
text list "SDC_G120D": 0 ''; 0 'Antrieb hat keine Störung / kein Fehlercode'; 1000 'Softwarefehler intern'; 1001 'FloatingPoint Ausnahme'; 1002 'Softwarefehler intern'; 1003 'Quittungsverzug bei Speicherzugriff'; 1004 'Softwarefehler intern'; 1005 'Datei Upload/Download fehlgeschlagen'; 1009 'CU: Regelungsbaugruppe Übertemperatur'; 1010 'Antriebstyp unbekannt'; 1015 'Softwarefehler intern'; 1016 'Firmware verändert'; 1017 'Komponentenlisten verändert'; 1018 'Hochlauf mehrmals abgebrochen'; 1019 'Wechselmedium schreiben fehlgeschlagen'; 1020 'RAM disk Schreiben fehlgeschlagen'; 1021 'Wechselmedium als USB-Datenträger von PC verwendet'; 1023 'Software Timeout intern'; 1028 'Konfigurationsfehler'; 1030 'Lebenszeichenausfall bei Steuerungshoheit'; 1033 'Einheitenumschaltung: Bezugsparameterwert ungültig'; 1034 'Einheitenumschaltung: Berechnung Parameterwerte nach Bezugswertänderung fehlgeschlagen'; 1035 'ACX: Parametersicherungsdateien beschädigt'; 1036 'ACX: Parametersicherungsdatei fehlt'; 1038 'ACX: Parametersicherungsdatei laden fehlgeschlagen'; 1039 'ACX: Parametersicherungsdatei schreiben fehlgeschlagen'; 1040 'Parameter sichern und POWER ON erforderlich'; 1042 'Parameterfehler beim Projekt-Download'; 1043 'Schwerer Fehler beim Projekt-Download'; 1044 'CU: Beschreibungsdaten fehlerhaft'; 1045 'Projektierungsdaten ungültig'; 1049 'Schreiben in Datei nicht möglich'; 1054 'CU: Systemgrenze überschritten'; 1064 'CU: Interner Fehler (CRC)'; 1066 'Zwischenspeicher: Füllstand 70 % erreicht oder überschritten'; 1067 'Zwischenspeicher: Füllstand 100 % erreicht'; 1068 'CU: Datenspeicher Speicherüberlauf'; 1069 'Parametersicherung und Gerät inkompatibel'; 1072 'Speicherkarte aus Sicherungskopie wieder hergestellt'; 1073 'POWER ON für Sicherungskopie auf Speicherkarte erforderlich'; 1105 'CU: Speicher nicht ausreichend'; 1107 'Speichern auf Speicherkarte fehlgeschlagen'; 1112 'CU: Leistungsteil unzulässig'; 1120 'Initialisierung Klemmen fehlgeschlagen'; 1122 'Frequenz am Messtastereingang zu hoch'; 1205 'CU: Zeitscheibenüberlauf'; 1250 'CU: CU-EEPROM Read-Only-Daten fehlerhaft'; 1251 'CU: CU-EEPROM Read-Write-Daten fehlerhaft'; 1257 'CU: Firmware-Version veraltet'; 1340 'Topologie: Zu viele Komponenten an einem Strang'; 1505 'BICO: Verschaltung kann nicht hergestellt werden'; 1510 'BICO: Signalquelle ist nicht Float'; 1511 'BICO: Verschaltung mit unterschiedlicher Normierung'; 1512 'BICO: Keine Normierung vorhanden'; 1513 'BICO: Verschaltung DO-übergreifend mit unterschiedlicher Normierung'; 1514 'BICO: Fehler beim Schreiben während Reconnect'; 1515 'BICO: Parameterschreiben nicht erlaubt da Steuerungshoheit aktiv'; 1590 'Antrieb: Motor Wartungsintervall abgelaufen'; 1600 'SI P1: STOP A ausgelöst'; 1611 'SI P1: Defekt in einem Überwachungskanal'; 1620 'SI P1: Sicher abgeschaltetes Moment aktiv'; 1625 'SI P1: Lebenszeichen in Safety-Daten fehlerhaft'; 1649 'SI P1: Softwarefehler intern'; 1650 'SI P1: Abnahmetest erforderlich'; 1651 'SI P1: Synchronisation Safety-Zeitscheiben fehlgeschlagen'; 1653 'SI P1: PROFIBUS/PROFINET-Projektierung fehlerhaft'; 1654 'SI P1: PROFIsafe-Projektierung abweichend'; 1655 'SI P1: Abgleich der Überwachungsfunktionen'; 1656 'SI P1: Parameter Prozessor 2 fehlerhaft'; 1658 'SI P1: PROFIsafe-Telegrammnummer ungeeignet'; 1659 'SI P1: Schreibauftrag für Parameter abgewiesen'; 1660 'SI P1: Sichere Funktionen nicht unterstützt'; 1661 'SI P1: Simulation der Safety Eingänge aktiv'; 1662 'Fehler interne Kommunikation'; 1663 'SI P1: Kopieren der SI-Parameter abgelehnt'; 1665 'SI P1: System ist defekt'; 1666 'SI Motion P1: Statisches 1-Signal am F-DI für sichere Quittierung'; 1669 'SI Motion: Kombination von Motor und Leistungsteil ungünstig'; 1680 'SI Motion P1: Prüfsummenfehler sichere Überwachungen'; 1681 'SI Motion P1: Parameterwert falsch'; 1682 'SI Motion P1: Überwachungsfunktion nicht unterstützt'; 1683 'SI Motion P1: SLS-Freigabe fehlt'; 1690 'SI Motion: Datensicherungsproblem beim NVRAM'; 1692 'SI Motion P1: Parameterwert geberlos unzulässig'; 1693 'SI Motion P1: Safety-Parametrierung geändert POWER ON erforderlich'; 1696 'SI Motion: Testanwahl der Bewegungsüberwachungen im Hochlauf'; 1697 'SI Motion: Test der Bewegungsüberwachungen erforderlich'; 1698 'SI P1: Inbetriebnahmemodus aktiv'; 1699 'SI P1: Test der Abschaltpfade erforderlich'; 1700 'SI Motion P1: STOP A ausgelöst'; 1701 'SI Motion P1: STOP B ausgelöst'; 1706 'SI Motion P1: SAM/SBR Grenze überschritten'; 1711 'SI Motion P1: Defekt in einem Überwachungskanal'; 1712 'SI Motion P1: Defekt bei F-IO-Verarbeitung'; 1714 'SI Motion P1: Sicher begrenzte Geschwindigkeit überschritten'; 1716 'SI Motion P1: Toleranz für sichere Bewegungsrichtung überschritten'; 1770 'SI Motion P1: Diskrepanzfehler der fehlersicheren Eingänge'; 1772 'SI Motion P1: Teststop fehlersichere Eingänge/Ausgänge aktiv'; 1773 'SI Motion P1: Teststop fehlerhaft'; 1774 'SI Motion P1: Teststop notwendig'; 1796 'SI P1: Warten auf Kommunikation'; 1798 'SI Motion P1: Teststop läuft'; 1799 'SI Motion P1: Abnahmetestmodus aktiv'; 1900 'PROFIBUS: Konfigurationstelegramm fehlerhaft'; 1910 'Feldbus SS Sollwert Timeout'; 1920 'PROFIBUS: Unterbrechung zyklische Verbindung'; 1945 'PROFIBUS: Verbindung zum Publisher gestört'; 1946 'PROFIBUS: Verbindung zum Publisher abgebrochen'; 1951 'CU SYNC: Synchronisation Applikationstakt fehlt'; 1953 'CU SYNC: Synchronisation nicht abgeschlossen'; 2050 'Trace: Start nicht möglich'; 2055 'Trace: Aufzeichnungsdauer zu klein'; 2056 'Trace: Aufzeichnungstakt zu klein'; 2057 'Trace: Zeitscheibentakt ungültig'; 2058 'Trace: Zeitscheibentakt für Endlostrace ungültig'; 2059 'Trace: Zeitscheibentakt für 2 x 8 Aufzeichnungskanäle ungültig'; 2060 'Trace: Aufzuzeichnendes Signal fehlt'; 2061 'Trace: Signal ungültig'; 2062 'Trace: Triggersignal ungültig'; 2063 'Trace: Datentyp ungültig'; 2070 'Trace: Parameter nicht änderbar'; 2075 'Trace: Pretriggerzeit zu groß'; 2080 'Trace: Parametrierung wegen Einheitenumschaltung gelöscht'; 2097 'MTrace: Mehrfachtrace aktivieren nicht möglich'; 2098 'MTrace: Speichern nicht möglich'; 2099 'Trace: Speicherplatz der Control Unit nicht ausreichend'; 2150 'OA: Applikation nicht ladbar'; 2151 'OA: Softwarefehler intern'; 2152 'OA: Speicher nicht ausreichend'; 3000 'NVRAM Fehler bei Aktion'; 3001 'NVRAM Prüfsumme fehlerhaft'; 3505 'CU: Analogeingang Drahtbruch'; 3510 'CU: Kalibrierdaten nicht plausibel'; 5000 'Leistungsteil: Übertemperatur Kühlkörper Wechselrichter'; 5001 'Leistungsteil: Übertemperatur Sperrschicht Chip'; 5002 'Leistungsteil: Übertemperatur Zuluft'; 5004 'Leistungsteil: Übertemperatur Gleichrichter'; 5006 'Leistungsteil: Übertemperatur Thermisches Modell'; 6310 'Anschlussspannung (p0210) fehlerhaft parametriert'; 6921 'Bremswiderstand Phasenunsymmetrie'; 6922 'Bremswiderstand Phasenausfall'; 7011 'Antrieb: Motor Übertemperatur'; 7012 'Antrieb: Motortemperaturmodell 1 Übertemperatur'; 7014 'Antrieb: Motortemperaturmodell Konfiguration Warnung'; 7015 'Antrieb: Motortemperatursensor Warnung'; 7016 'Antrieb: Motortemperatursensor Störung'; 7080 'Antrieb: Regelungsparameter fehlerhaft'; 7082 'Makro: Ausführung nicht möglich'; 7083 'Makro: ACX-File nicht gefunden'; 7084 'Makro: Bedingung für WaitUntil nicht erfüllt'; 7086 'Einheitenumschaltung: Parametergrenzverletzung durch Bezugswertänderung'; 7088 'Einheitenumschaltung: Parametergrenzverletzung durch Einheitenumschaltung'; 7089 'Einheitenumschaltung: Funktionsmodul aktivieren ist blockiert weil Einheiten umgeschaltet'; 7200 'Antrieb: Steuerungshoheit EIN-Befehl steht an'; 7220 'Antrieb: Führung durch PLC fehlt'; 7300 'Antrieb: Netzschütz Rückmeldung fehlt'; 7320 'Antrieb: Automatischer Wiederanlauf abgebrochen'; 7321 'Antrieb: Automatischer Wiederanlauf aktiv'; 7330 'Fangen: Gemessener Suchstrom zu klein'; 7331 'Fangen: Funktion nicht unterstützt'; 7400 'Antrieb: Zwischenkreisspannungs-Maximum-Regler aktiv'; 7401 'Antrieb: Zwischenkreisspannungs-Maximum-Regler deaktiviert'; 7402 'Antrieb: Zwischenkreisspannungs-Minimum-Regler aktiv'; 7404 'Antrieb: Zwischenkreisspannungsüberwachnung Vdc_Max'; 7405 'Antrieb: Kinetische Pufferung minimale Drehzahl unterschritten'; 7406 'Antrieb: Kinetische Pufferung maximale Dauer überschritten'; 7409 'Antrieb: U/f-Steuerung Strombegrenzungsregler aktiv'; 7410 'Antrieb: Stromreglerausgang begrenzt'; 7411 'Antrieb: Flussreglerausgang begrenzt'; 7416 'Antrieb: Konfiguration Flussregler'; 7426 'Technologieregler Istwert begrenzt'; 7428 'Technologieregler Parametrierfehler'; 7435 'Antrieb: Hochlaufgebersetzen bei geberloser Vektorregelung'; 7440 'EPOS: Ruckzeit wird begrenzt'; 7441 'LR: Lageoffset der Absolutwertgeberjustage sichern'; 7442 'LR: Multiturn passt nicht zum Modulobereich'; 7443 'LR: Referenzpunkt-Koordinate nicht im zulässigen Bereich'; 7450 'LR: Stillstandsüberwachung hat angesprochen'; 7451 'LR: Positionierüberwachung hat angesprochen'; 7452 'LR: Schleppabstand zu groß'; 7453 'LR: Lageistwertaufbereitung fehlerhaft'; 7454 'LR: Lageistwertaufbereitung hat keinen gültigen Geber'; 7455 'EPOS: Maximalgeschwindigkeit begrenzt'; 7456 'EPOS: Sollgeschwindigkeit begrenzt'; 7457 'EPOS: Eingangssignale Kombination unzulässig'; 7458 'EPOS: Referenznocken nicht gefunden'; 7459 'EPOS: Keine Nullmarke vorhanden'; 7460 'EPOS: Referenznockenende nicht gefunden'; 7461 'EPOS: Referenzpunkt nicht gesetzt'; 7462 'EPOS: Angewählte Verfahrsatznummer existiert nicht'; 7463 'EPOS: Externer Satzwechsel im Verfahrsatz nicht angefordert'; 7464 'EPOS: Verfahrsatz ist inkonsistent'; 7465 'EPOS: Verfahrsatz hat keinen Folgesatz'; 7466 'EPOS: Verfahrsatznummer mehrfach vergeben'; 7467 'EPOS: Verfahrsatz hat unzulässigen Auftragsparameter'; 7468 'EPOS: Verfahrsatz Sprungziel existiert nicht'; 7469 'EPOS: Verfahrsatz Zielposition < Software-Endschalter Minus'; 7470 'EPOS: Verfahrsatz Zielposition > Software-Endschalter Plus'; 7471 'EPOS: Verfahrsatz Zielposition außerhalb Modulobereich'; 7472 'EPOS: Verfahrsatz ABS_POS/ABS_NEG nicht möglich'; 7473 'EPOS: Verfahrbereichsanfang angefahren'; 7474 'EPOS: Verfahrbereichsende angefahren'; 7475 'EPOS: Zielposition < Verfahrbereichsanfang'; 7476 'EPOS: Zielposition > Verfahrbereichsende'; 7477 'EPOS: Zielposition < Software-Endschalter Minus'; 7478 'EPOS: Zielposition > Software-Endschalter Plus'; 7479 'EPOS: Software-Endschalter Minus angefahren'; 7480 'EPOS: Software-Endschalter Plus angefahren'; 7481 'EPOS: Achsposition < Software-Endschalter Minus'; 7482 'EPOS: Achsposition > Software-Endschalter Plus'; 7483 'EPOS: Fahren auf Festanschlag Klemmmoment nicht erreicht'; 7484 'EPOS: Festanschlag außerhalb Überwachungsfenster'; 7485 'EPOS: Festanschlag nicht erreicht'; 7486 'EPOS: Zwischenhalt fehlt'; 7487 'EPOS: Verfahrauftrag verwerfen fehlt'; 7488 'EPOS: Relative Positionierung nicht möglich'; 7489 'EPOS: Referenzpunktkorrektur außerhalb Fenster'; 7490 'EPOS: Freigabe während Verfahren weggenommen'; 7491 'EPOS: STOP-Nocken Minus angefahren'; 7492 'EPOS: STOP-Nocken Plus angefahren'; 7493 'LR: Überlauf des Wertebereiches für Lageistwert'; 7494 'LR: Antriebsdatensatz-Umschaltung während Betrieb'; 7495 'LR: Referenzfunktion abgebrochen'; 7496 'EPOS: Freigabe nicht möglich'; 7497 'LR: Lagesetzwert aktiviert'; 7498 'LR: Messtasterauswertung nicht möglich'; 7499 'EPOS: Umkehrnocken mit falscher Verfahrrichtung angefahren'; 7503 'EPOS: STOP-Nocken mit falscher Verfahrrichtung angefahren'; 7505 'EPOS: Auftrag Festanschlag bei U/f/SLVC-Betrieb nicht möglich'; 7530 'Antrieb: Antriebsdatensatz DDS nicht vorhanden'; 7531 'Antrieb: Befehlsdatensatz CDS nicht vorhanden'; 7550 'Antrieb: Geberparameter zurücksetzen nicht möglich'; 7552 'Antrieb Geber: Geberkonfiguration nicht unterstützt'; 7553 'Antrieb Geber: Sensor Module Konfiguration nicht unterstützt'; 7557 'Geber 1: Referenzpunkt-Koordinate nicht im zulässigen Bereich'; 7558 'Geber 2: Referenzpunkt-Koordinate nicht im zulässigen Bereich'; 7563 'Antrieb Geber: XIST1_ERW Konfiguration fehlerhaft'; 7565 'Antrieb: Geberfehler PROFIdrive-Geberschnittstelle 1'; 7566 'Antrieb: Geberfehler PROFIdrive-Geberschnittstelle 2'; 7577 'Geber 1: Messtasterauswertung nicht möglich'; 7578 'Geber 2: Messtasterauswertung nicht möglich'; 7581 'Geber 1: Lageistwertaufbereitung fehlerhaft'; 7582 'Geber 2: Lageistwertaufbereitung fehlerhaft'; 7584 'Geber 1: Lagesetzwert aktiviert'; 7585 'Geber 2: Lagesetzwert aktiviert'; 7587 'Geber 1: Lageistwertaufbereitung hat keinen gültigen Geber'; 7588 'Geber 2: Lageistwertaufbereitung hat keinen gültigen Geber'; 7590 'Geber 1: Antriebsdatensatz-Umschaltung während Betrieb'; 7591 'Geber 2: Antriebsdatensatz-Umschaltung während Betrieb'; 7593 'Geber 1: Wertebereich für Lageistwert überschritten'; 7594 'Geber 2: Wertebereich für Lageistwert überschritten'; 7596 'Geber 1: Referenzfunktion abgebrochen'; 7597 'Geber 2: Referenzfunktion abgebrochen'; 7599 'Geber 1: Justage nicht möglich'; 7600 'Geber 2: Justage nicht möglich'; 7800 'Antrieb: Kein Leistungsteil vorhanden'; 7801 'Antrieb: Motor Überstrom'; 7802 'Antrieb: Einspeisung oder Leistungsteil nicht bereit'; 7805 'Antrieb: Leistungsteil Überlastung I2t'; 7806 'Antrieb: Generatorische Leistungsgrenze überschritten (F3E)'; 7807 'Antrieb: Kurzschluss/Erdschluss erkannt'; 7808 'HF Damping Module: Dämpfung nicht bereit'; 7810 'Antrieb: Leistungsteil-EEPROM ohne Nenndaten'; 7850 'Externe Warnung 1'; 7851 'Externe Warnung 2'; 7852 'Externe Warnung 3'; 7860 'Externe Störung 1'; 7861 'Externe Störung 2'; 7862 'Externe Störung 3'; 7900 'Antrieb: Motor blockiert'; 7901 'Antrieb: Motor Überdrehzahl'; 7902 'Antrieb: Motor gekippt'; 7903 'Antrieb: Motor Drehzahlabweichung'; 7910 'Antrieb: Motor Übertemperatur'; 7920 'Antrieb: Drehmoment/Drehzahl zu niedrig'; 7921 'Antrieb: Drehmoment/Drehzahl zu hoch'; 7922 'Antrieb: Drehmoment/Drehzahl außerhalb Toleranz'; 7923 'Antrieb: Drehmoment/Drehzahl zu niedrig'; 7924 'Antrieb: Drehmoment/Drehzahl zu hoch'; 7925 'Antrieb: Drehmoment/Drehzahl außerhalb Toleranz'; 7927 'Gleichstrombremsung aktiv'; 7929 'Antrieb: Kein Motor erkannt'; 7936 'Antrieb: Lastausfall'; 7950 'Motorparameter fehlerhaft'; 7967 'Antrieb: Pollageidentifikation interner Fehler'; 7968 'Antrieb: Lq-Ld-Messung fehlerhaft'; 7969 'Antrieb: Pollageidentifikation fehlerhaft'; 7975 'Antrieb: Fahren bis Nullmarke - Sollwertvorgabe erwartet'; 7976 'Antrieb: Geberfeinabgleich aktiviert'; 7980 'Antrieb: Drehende Messung aktiviert'; 7981 'Antrieb: Drehende Messung Freigaben fehlen'; 7983 'Antrieb: Drehende Messung Sättigungskennlinie'; 7984 'Antrieb: Drehzahlregleroptimierung Trägheitsmoment'; 7985 'Antrieb: Drehzahlregleroptimierung (Schwingungstest)'; 7986 'Antrieb: Drehende Messung Hochlaufgeber'; 7988 'Antrieb: Drehende Messung Keine Konfiguration ausgewählt'; 7990 'Antrieb: Motordatenidentifikation fehlerhaft'; 7991 'Antrieb: Motordatenidentifikation aktiviert'; 7994 'Antrieb: Motordatenidentifikation nicht durchgeführt'; 8010 'CU: Analog-Digital-Wandler'; 8501 'PROFINET: Sollwert Timeout'; 8502 'PROFINET: Überwachungszeit Lebenszeichen abgelaufen'; 8511 'PROFINET: Empfangs-Konfigurationsdaten ungültig'; 8526 'PROFINET: Keine zyklische Verbindung'; 8565 'PROFINET: Konsistenzfehler bei Einstellparametern'; 8760 'CAN: Überschreitung maximaler Größe des PZD IF'; 8800 'PROFIenergy Energiesparmodus aktiv'; 8802 'PROFIenergy Inkrementalgeberversorgung ausschalten nicht möglich'; 13009 'Lizenzierung OA-Applikation nicht lizenziert'; 13100 'Know-how-Schutz: Kopierschutzfehler'; 13101 'Know-how-Schutz: Kopierschutz nicht aktivierbar'; 13102 'Know-how-Schutz: Konsistenzfehler der geschützten Daten'; 30001 'Leistungsteil: Überstrom'; 30002 'Leistungsteil: Zwischenkreisspannung Überspannung'; 30003 'Leistungsteil: Zwischenkreisspannung Unterspannung'; 30004 'Leistungsteil: Übertemperatur Kühlkörper Wechselrichter'; 30005 'Leistungsteil: Überlastung I2t'; 30011 'Leistungsteil: Netzphasenausfall im Hauptstromkreis'; 30015 'Leistungsteil: Phasenausfall Motorleitung'; 30016 'Leistungsteil: Lastversorgung ausgeschaltet'; 30017 'Leistungsteil: Hardware Strombegrenzung zu oft angesprochen'; 30021 'Leistungsteil: Erdschluss'; 30022 'Leistungsteil: Überwachung U_ce'; 30024 'Leistungsteil: Übertemperatur Thermisches Modell'; 30025 'Leistungsteil: Übertemperatur Chip'; 30027 'Leistungsteil: Vorladung Zwischenkreis Zeitüberwachung'; 30031 'Leistungsteil: Hardware Strombegrenzung in Phase U'; 30032 'Leistungsteil: Hardware Strombegrenzung in Phase V'; 30033 'Leistungsteil: Hardware Strombegrenzung in Phase W'; 30034 'Leistungsteil: Übertemperatur Innenraum'; 30042 'Leistungsteil: Lüfter hat maximale Betriebsstunden erreicht'; 30052 'EEPROM Daten fehlerhaft'; 30054 'Leistungsteil: Unterspannung bei Bremse öffnen'; 30057 'Leistungsteil: Netzunsymmetrie'; 30071 'Keine neuen Istwerte von Power Module empfangen'; 30072 'Keine Sollwerte mehr an Power Module übertragbar'; 30074 'Kommunikationsfehler zwischen Control Unit und Power Module'; 30080 'Leistungsteil: Stromanstieg zu schnell'; 30081 'Leistungsteil: Schalthandlungen zu häufig'; 30105 'LT: Istwerterfassung fehlerhaft'; 30502 'Leistungsteil: Zwischenkreis Überspannung'; 30600 'SI P2: STOP A ausgelöst'; 30611 'SI P2: Defekt in einem Überwachungskanal'; 30620 'SI P2: Sicher abgeschaltetes Moment aktiv'; 30625 'SI P2: Lebenszeichen in Safety-Daten fehlerhaft'; 30649 'SI P2: Softwarefehler intern'; 30650 'SI P2: Abnahmetest erforderlich'; 30651 'SI P2: Synchronisation mit Control Unit fehlgeschlagen'; 30655 'SI P2: Abgleich der Überwachungsfunktionen'; 30656 'SI P2: Parameter Prozessor 2 fehlerhaft'; 30659 'SI P2: Schreibauftrag für Parameter abgewiesen'; 30662 'Fehler in interner Kommunikation'; 30664 'Fehler in der Hochlaufphase'; 30665 'SI P2: System ist defekt'; 30666 'SI Motion P2: Statisches 1-Signal am F-DI für sichere Quittierung'; 30680 'SI Motion P2: Prüfsummenfehler sichere Überwachungen'; 30681 'SI Motion P2: Parameterwert falsch'; 30682 'SI Motion P2: Überwachungsfunktion nicht unterstützt'; 30683 'SI Motion P2: SLS-Freigabe fehlt'; 30692 'SI Motion P2: Parameterwert falsch geberlos'; 30693 'SI P2: Safety-Parametrierung geändert POWER ON erforderlich'; 30700 'SI Motion P2: STOP A ausgelöst'; 30701 'SI Motion P2: STOP B ausgelöst'; 30706 'SI Motion P2: SAM/SBR Grenze überschritten'; 30711 'SI Motion P2: Defekt in einem Überwachungskanal'; 30712 'SI Motion P2: Defekt bei F-IO-Verarbeitung'; 30714 'SI Motion P2: Sicher begrenzte Geschwindigkeit überschritten'; 30716 'SI Motion P2: Toleranz für sichere Bewegungsrichtung überschritten'; 30770 'SI Motion P2: Diskrepanzfehler der fehlersicheren Eingänge'; 30772 'SI Motion P2: Teststop fehlersichere Eingänge/Ausgänge aktiv'; 30773 'SI Motion P2: Teststop fehlerhaft'; 30798 'SI Motion P2: Teststop läuft'; 30799 'SI Motion P2: Abnahmetestmodus aktiv'; 30800 'Leistungsteil: Sammelmeldung'; 30802 'Leistungsteil: Zeitscheibenüberlauf'; 30804 'Leistungsteil: CRC'; 30805 'Leistungsteil: Prüfsumme EPROM nicht korrekt'; 30809 'Leistungsteil: Schaltinformation ungültig'; 30810 'Leistungsteil: Watchdog Timer'; 30850 'Leistungsteil: Softwarefehler intern'; 30875 'Leistungsteil DRIVE-CLiQ (CU): Versorgungsspannung ausgefallen'; 30903 'Leistungsteil: I2C-Bus Fehler aufgetreten'; 30920 'Fehler Temperatursensor'; 30950 'Leistungsteil: Softwarefehler intern'; 30999 'Leistungsteil: Unbekannte Warnung'; 31100 'Geber 1: Nullmarkenabstand fehlerhaft'; 31101 'Geber 1: Nullmarke ausgefallen'; 31103 'Geber 1: Amplitudenfehler Spur R'; 31118 'Geber 1: Drehzahldifferenz außerhalb Toleranz'; 31131 'Geber 1: Abweichung Lage inkrementell/absolut zu groß'; 31150 'Geber 1: Initialisierung fehlerhaft'; 31400 'Geber 1: Warnschwelle Nullmarkenabstand fehlerhaft'; 31401 'Geber 1: Warnschwelle Nullmarke ausgefallen'; 31418 'Geber 1: Drehzahldifferenz je Abtastrate überschritten'; 31422 'Geber 1: Impulszahl Rechteckgeber außerhalb Toleranzband'; 31431 'Geber 1: Abweichung Lage inkrementell/absolut zu groß'; 31802 'Geber 1: Zeitscheibenüberlauf'; 31805 'Geber 1: Prüfsumme EPROM nicht korrekt'; 31850 'Geber 1: Geberauswertung Softwarefehler intern'; 31899 'Geber 1: Unbekannte Störung'; 31905 'Geber 1: Fehlparametrierung'; 31915 'Geber 1: Konfigurationsfehler'; 31930 'Geber 1: Datalogger hat Daten gespeichert'; 31950 'Geber 1: Softwarefehler intern'; 31999 'Geber 1: Unbekannte Warnung'; 32110 'Geber 2: Serielle Kommunikation gestört'; 32111 'Geber 2: Absolutwertgeber interner Fehler'; 32112 'Geber 2: Fehlerbit im seriellen Protokoll gesetzt'; 32150 'Geber 2: Initialisierung fehlerhaft'; 32410 'Geber 2: Serielle Kommunikation'; 32411 'Geber 2: Absolutwertgeber meldet Warnungen'; 32412 'Geber 2: Fehlerbit im seriellen Protokoll gesetzt'; 32442 'Geber 2: Batteriespannung Vorwarnung'; 32802 'Geber 2: Zeitscheibenüberlauf'; 32805 'Geber 2: Prüfsumme EPROM nicht korrekt'; 32850 'Geber 2: Geberauswertung Softwarefehler intern'; 32899 'Geber 2: Unbekannte Störung'; 32905 'Geber 2: Fehlparametrierung'; 32915 'Geber 2: Konfigurationsfehler'; 32930 'Geber 2: Datalogger hat Daten gespeichert'; 32950 'Geber 2: Softwarefehler intern'; 32999 'Geber 2: Unbekannte Warnung'; 50001 'PROFINET Konfigurationsfehler'; 50010 'PROFINET Name of Station ungültig'; 50020 'PROFINET: Zweiter Controller fehlt'; 50510 'FBLOCKS: Anmeldung der Ablaufgruppe abgelehnt'; 50511 'FBLOCKS: Kein Speicher für Freie Funktionsblöcke mehr verfügbar'; 50513 'FBLOCKS: Ablaufreihenfolgewert bereits vergeben'; 50517 'FBLOCKS: Interne Messung aktiv'; 50518 'FBLOCKS: Abtastzeit freie Ablaufgruppe weicht bei Downloaden ab'; 30051 'Leistungsteil: Motorhaltebremse Kurzschluss erkannt'

text list "SDC_ScreensName": 0 '---'; 100 'SDC - Diagnose PN: / Diagnostics Overview SDC PN:'; 101 'SDC - Diagnose PN: / Diagnostics Overview SDC PN:'; 160 'SDC - HOME / Start'; 700 'SDC - global parameter / Global Parameter'; 703 'SDC - barcode jumps / Barcode Leaps / Barcode Sprünge'; 704 'SDC - TS parameter drive / TS Parameter Drive'; 705 'SDC - TS parameter hoist / TS Parameter Hoist'; 711 'SDC - EMS status / EMS Status'; 724 'SDC - error archiv / Fault Status Archiev / Error History'; 726 'SDC - EMS Simulation / EMS Simulation'; 734 'SDC - barcode inserts / Barcode Inserts/Cuts / Barcode Missions/Cuts Correction Table'; 735 'SDC - distance control snychron area / Distance Control Snychron Area / Distance Control Synchron Area'; 736 'SDC - distance control limits / Distance Control Limits not in snychron Area / Distance Control Limits not in synchron Area'; 161 'SDC - plant overview brown field 1 / Overview'; 190 'SDC - errors / Messages'; 701 'SDC - EMS Flags / EMS Flags'; 728 'SDC - EMS status G120D / EMS Status G120D'; 712 'SDC - EMS status I/O / EMS Status / EMS Status IO'; 702 'SDC - EMS parameter'; 7020 'SDC - EMS parameter drive'; 7021 'SDC - EMS parameter hoist'; 722 'SDC - EMS errors'; 716 'SDC - track section status / TS IF'; 162 'SDC - plant overview brown field 2 / Overview'; 163 'SDC - plant overview green field'; 752 'Profinet Diagnostics'

text list "SDC_ER_EMS": 501 'Error emergency stop / Störung Not Halt / Error Not Halt'; 502 'Error Fuse 000EEA001FC2 (+24V) / Störung Sicherung BS1FC302 / Error Sicherung F2'; 503 'Error VAC ID / Störung EMS ID / Error EMS ID'; 504 'Error heartbeat / Störung Lebensbit / Error Lebensbit'; 505 'Error Safety-Module KFA001.2 fault (cabinet) / Störung Safety-Modul KFA131 gestört (Schaltkasten) / Error Safety-Modul KFA131 gestört (Schaltkasten)'; 506 'Error Safety-Module KFA001.3 fault (cabinet) / Reserve'; 507 'Error Safety-Module KFA001.4 fault (cabinet) / Störung Safety-Modul KFA141 gestört (Schaltkasten) / Error Safety-Modul KFA141 gestört (Schaltkasten)'; 508 'Error Fuse 000AKL001QA1 (480V Deutronic) / Reserve'; 509 'Error Profinet trolly-FI -TA005 / Störung Profinet Fahr-FU FE1TA1 / Error Profinet Fahr-FU'; 510 'Error Profinet hoist-FI -TA006 / Störung Profinet Hub-FU HE1TA1 / Error Profinet Hub-FU'; 511 'Error Profinet Scanner Leutze -KG004 / Störung Profinet AposOptic 1 FE1BX01 / Error Profinet Scanner 1'; 512 'spare / Störung Profinet AposOptic 2 FE1BX02 / Error Profinet Scanner 2'; 513 'Error Profinet hoist rope encoder -GF003 / Störung Profinet Hub Seilgeber HE1GF1 / Error Profinet Hub Seilgeber'; 514 'spare / Reserve'; 515 'Error Profinet Error WiFi Client / Störung Kommunikationsmodul BS1TFC1 / Error Kommunikationsmodul'; 516 'spare / Reserve'; 517 'Error Deutronic / Störung Profinet Schwenk Drehgeber (T&R) SN1GF1 / Error Profinet Schwenk Drehgeber (T&R)'; 518 'Error Profinet: spare / Reserve'; 519 'Error Profinet: spare / Reserve'; 520 'Error Profinet: spare / Reserve'; 521 'Error Profinet: spare / Reserve'; 522 'Error Profinet: spare / Reserve'; 523 'Error Profinet: spare / Reserve'; 524 'Error Profinet: spare / Reserve'; 525 'Error Safety-Module -TA005 fault (trolly-FI) / Störung Safety-Modul FE1TA1 gestört (Fahr-FU) / Error Safety-Modul TA1 gestört (Fahr-FU)'; 526 'Error Safety-Module -TA006 fault (hoist-FI) / Störung Safety-Modul HE1TA1 gestört (Hub-FU) / Error Safety-Modul TA2 gestört (Hub-FU)'; 527 'Error Deutronic invalid feedback / Störung Safety-Modul SN1TA1 gestört (Schwenk-FU) / Error Safety-Modul TA3 gestört (Schwenk-FU)'; 528 'spare / Reserve'; 529 'spare / Reserve'; 530 'spare / Reserve'; 531 'spare / Reserve'; 532 'Error PLC / Störung SPS'; 801 'Warning no feedback vacuum cleaner / Meldung keine Rückmeldung Staubsauger / Reserve'; 802 'Warning motor protection circuit breake vacuum cleaner / Meldung Motorschutz Staubsauger / Reserve'; 803 'Warning Deutronic device error / Reserve'; 804 'Warning Deutronic handling error / Reserve'; 805 'warning spare / Reserve'; 806 'warning spare / Reserve'; 807 'warning spare / Reserve'; 808 'warning spare / Reserve'; 809 'warning spare / Reserve'; 810 'warning spare / Reserve'; 811 'warning spare / Reserve'; 812 'warning spare / Reserve'; 813 'warning spare / Reserve'; 814 'warning spare / Reserve'; 815 'warning spare / Reserve'; 816 'warning spare / Reserve'; 817 'Warning bypass active / Meldung Bypass eingeschaltet / Anzeige Bypass eingeschaltet'; 818 'Warning Initialization hoist / Meldung Initialisierung Hub / Anzeige Initialisierung Hub'; 819 'warning spare / Reserve / Anzeige Störung von SDC liegt vor'; 820 'warning spare / Reserve / Anzeige Download FU-Parameter läuft'; 821 'warning spare / Reserve / Anzeige Fangbremse und Schalter prüfen'; 822 'Warning VAC IR manual operation activated / Reserve'; 823 'Warning SDC manual operation activated / Meldung SDC hat Betriebsart Hand angewählt / Anzeige SDC hat Betriebsart Hand angewählt'; 824 'Warning Emergency Stop in track section / Meldung NotAus von Anlagen-SPS / Anzeige NotAus von Anlagen-SPS'; 825 'Warning distance control / Meldung Distanzkontrolle / Anzeige Distanzkontrolle'; 826 'warning EMS in manual mode / Reserve'; 827 'warning spare / Reserve'; 828 'Warning emergency mode drive unit active / Meldung Notbetrieb ein Fahrantrieb angewählt / Anzeige Notbetrieb ein Hubantrieb angewählt'; 829 'warning spare / Meldung Notbetrieb ein Schwenkantrieb angewählt / Anzeige Notbetrieb ein Schwenkantrieb angewählt'; 830 'Warning emergency mode hoist unit active / Meldung Notbetrieb ohne Hub angewählt / Anzeige Notbetrieb ohne Hub angewählt'; 831 'warning spare / Reserve'; 832 'warning spare / Reserve'; 601 'Error trolley: frequency inverter / Störung Fahrantrieb: Frequenzumrichter / Error Drive: Frequenzumrichter'; 602 'spare / Reserve / Fault Drive Scanner: 24V DC'; 603 'Error trolley: drive command not plausible / Störung Fahrantrieb: Antriebskommando nicht plausibel / Error Drive: Antriebskommando nicht plausibel'; 604 'spare / Reserve / Fault Drive Scanner: 24V DC'; 605 'Error trolley: scanner invalid value / Reserve / Fault Drive Scanner: 24V DC'; 606 'spare / Reserve / Fault Drive Scanner: 24V DC'; 607 'Error trolley: speed too high / Störung Fahrantrieb: Geschwindigkeit zu hoch / Error Drive: Geschwindigkeit zu hoch'; 608 'Error trolley: speed too low / Störung Fahrantrieb: Geschwindigkeit zu niedrig / Error Drive: Geschwindigkeit zu niedrig'; 609 'Error trolley: movement without enable / Störung Fahrantrieb: Bewegung ohne Freigabe / Error Drive: Bewegung ohne Freigabe'; 610 'Error trolley: positioning - jump not plausible / Störung Fahrantrieb: Positionserkennung: Sprung unzulässig / Error Drive Scanner: Sprung unzulässig'; 611 'Error trolley: setpoint passed / Störung Fahrantrieb: Positionierpunkt überfahren / Fault Drive Stop position overrun'; 612 'Error trolley: no valid scanner value (quality) / Reserve / Fault Drive Scanner: 24V DC'; 613 'Error trolley: spare / Reserve / Fault Drive Scanner: 24V DC'; 614 'Error trolley: spare / Reserve / Fault Drive Scanner: 24V DC'; 615 'Error trolley: spare / Reserve / Fault Drive Scanner: 24V DC'; 616 'Error trolley: spare / Reserve / Fault Drive Scanner: 24V DC'; 617 'Error trolley: spare / Reserve / Fault Drive Scanner: 24V DC'; 618 'Error trolley: spare / Reserve / Fault Drive Scanner: 24V DC'; 619 'Error trolley: spare / Reserve / Fault Drive Scanner: 24V DC'; 620 'Error trolley: spare / Reserve / Fault Drive Scanner: 24V DC'; 621 'Error trolley: spare / Reserve / Fault Drive Scanner: 24V DC'; 622 'Error trolley: spare / Reserve / Fault Drive Scanner: 24V DC'; 623 'Error trolley: spare / Reserve / Fault Drive Scanner: 24V DC'; 624 'Error trolley: spare / Reserve / Fault Drive Scanner: 24V DC'; 625 'Error trolley: spare / Reserve / Fault Drive Scanner: 24V DC'; 626 'Error trolley: spare / Reserve / Fault Drive Scanner: 24V DC'; 627 'Error trolley: spare / Reserve / Fault Drive Scanner: 24V DC'; 628 'Error trolley: spare / Reserve / Fault Drive Scanner: 24V DC'; 629 'Error trolley: spare / Reserve / Fault Drive Scanner: 24V DC'; 630 'Error trolley: spare / Reserve / Fault Drive Scanner: 24V DC'; 631 'Error trolley: spare / Reserve / Fault Drive Scanner: 24V DC'; 632 'Error trolley: spare / Reserve / Fault Drive Scanner: 24V DC'; 633 'Error trolley FI: overcurrent / Störung Fahrantrieb FU 1: Überstrom / Error Drive FU 1: Überstrom'; 634 'Error trolley FI: DC bus voltage overvoltage / Störung Fahrantrieb FU 1: Zwischenkreisspannung Überspannung / Error Drive FU 1: Zwischenkreisspannung Überspannung'; 635 'Error trolley FI: DC bus voltage undervoltage / Störung Fahrantrieb FU 1: Zwischenkreisspannung Unterspannung / Error Drive FU 1: Zwischenkreisspannung Unterspannung'; 636 'Error trolley FI: overtemperature / Störung Fahrantrieb FU 1: Übertemperatur Kühlkörper Wechselrichter / Error Drive FU 1: Übertemperatur Kühlkörper Wechselrichter'; 637 'Error trolley FI: error on driver identification / Störung Fahrantrieb FU 1: Motordatenidentifikation fehlerhaft / Error Drive FU 1: Motordatenidentifikation fehlerhaft'; 638 'Error trolley FI: ground / Störung Fahrantrieb FU 1: Erdschluss / Error Drive FU 1: Erdschluss'; 639 'Error trolley: spare / Reserve / Fault Drive Scanner: 24V DC'; 640 'Error trolley FI: control requested from PLC / Störung Fahrantrieb FU 1: Führung durch PLC fehlt / Error Drive FU 1: Führung durch PLC fehlt'; 641 'Error trolley FI: drive overtemperature / Störung Fahrantrieb FU 1: Reserve / Error Drive FU 1: Reserve'; 642 'Error trolley: spare / Reserve / Fault Drive Scanner: 24V DC'; 643 'Error trolley: spare / Reserve / Fault Drive Scanner: 24V DC'; 644 'Error trolley: spare / Reserve / Fault Drive Scanner: 24V DC'; 645 'Error trolley: spare / Reserve / Fault Drive Scanner: 24V DC'; 646 'Error trolley: spare / Reserve / Fault Drive Scanner: 24V DC'; 647 'Error trolley: spare / Reserve / Fault Drive Scanner: 24V DC'; 648 'Error trolley: spare / Reserve / Fault Drive Scanner: 24V DC'; 649 'Error trolley Safety: scanner invalid jump / Störung Fahrantrieb Safety: AposOptic 1 Sprung nicht zulässig / Error Drive Safety: Scanner 1 Sprung nicht zulässig'; 650 'Error trolley Safety: G120D invalid jump / Störung Fahrantrieb Safety: AposOptic 2 Sprung nicht zulässig / Error Drive Safety: Scanner 2 Sprung nicht zulässig'; 651 'Error trolley Safety: Scanner limit exceeded / Störung Fahrantrieb Safety: AposOpticwert 1 hat Limit überschritten / Error Drive Safety: Scannerwert 1 hat Limit überschritten'; 652 'Error trolley Safety: G120D limit exceeded / Störung Fahrantrieb Safety: AposOpticwert 2 hat Limit überschritten / Error Drive Safety: Scannerwert 2 hat Limit überschritten'; 653 'Error trolley Safety: speed scanner to high / Störung Fahrantrieb Safety: Geschwindigkeit AposOpticwert 1 zu hoch / Error Drive Safety: Geschwindigkeit G120 Drehzahl zu hoch'; 654 'Error trolley Safety: value of scanner opposite to command / Störung Fahrantrieb Safety: Wertänderung des AposOpticwert 1 entspricht nicht der Drehrichtung / Error Drive Safety: Drehzahl des G120D entsprechen nicht der Drehrichtung'; 655 'Error trolley Safety: speed G120D to high / Störung Fahrantrieb Safety: Geschwindigkeit AposOpticwert 2 zu hoch / Error Drive Safety: Geschwindigkeit Barcode zu hoch'; 656 'Error trolley Safety: value of G120D opposite to command / Störung Fahrantrieb Safety: Wertänderung des AposOpticwert 2 entspricht nicht der Drehrichtung / Error Drive Safety: Wertänderung des Barcode entspricht nicht der Drehrichtung'; 657 'Error trolley Safety: Emergency Stop area not set / Störung Fahrantrieb Safety: Not Halt Bereich nicht deffiniert / Error Drive Safety: E-Stop Bereich nicht deffiniert'; 658 'Error trolley: spare / Reserve / Fault Drive Scanner: 24V DC'; 659 'Error trolley Safety: difference Scanner/G120D to high / Störung Fahrantrieb Safety: Differenz AposOptic 1 / 2 zu hoch / Error Drive Safety: Differenz Scanner 1 / 2 zu hoch'; 660 'Error trolley Safety: no enable of scanner / Störung Fahrantrieb Safety: Reserve / Error Drive Safety: Reserve'; 661 'Error trolley Safety: spare / Störung Fahrantrieb Safety: Reserve / Error Drive Safety: Reserve'; 662 'Error trolley Safety: spare / Störung Fahrantrieb Safety: Reserve / Error Drive Safety: Reserve'; 663 'Error trolley Safety: spare / Störung Fahrantrieb Safety: Reserve / Error Drive Safety: Reserve'; 664 'Error trolley Safety: spare / Störung Fahrantrieb Safety: Reserve / Error Drive Safety: Reserve'; 665 'spare / Störung Fahrantrieb FU 2: Überstrom / Error Drive FU 2: Überstrom'; 666 'spare / Störung Fahrantrieb FU 2: Überstrom / Error Drive FU 2: Überstrom'; 667 'spare / Störung Fahrantrieb FU 2: Überstrom / Error Drive FU 2: Überstrom'; 668 'spare / Störung Fahrantrieb FU 2: Überstrom / Error Drive FU 2: Überstrom'; 669 'spare / Störung Fahrantrieb FU 2: Überstrom / Error Drive FU 2: Überstrom'; 670 'spare / Störung Fahrantrieb FU 2: Überstrom / Error Drive FU 2: Überstrom'; 671 'spare / Störung Fahrantrieb FU 2: Überstrom / Error Drive FU 2: Überstrom'; 672 'spare / Störung Fahrantrieb FU 2: Überstrom / Error Drive FU 2: Überstrom'; 673 'spare / Störung Fahrantrieb FU 2: Überstrom / Error Drive FU 2: Überstrom'; 674 'spare / Störung Fahrantrieb FU 2: Überstrom / Error Drive FU 2: Überstrom'; 675 'spare / Störung Fahrantrieb FU 2: Überstrom / Error Drive FU 2: Überstrom'; 676 'spare / Störung Fahrantrieb FU 2: Überstrom / Error Drive FU 2: Überstrom'; 677 'spare / Störung Fahrantrieb FU 2: Überstrom / Error Drive FU 2: Überstrom'; 678 'spare / Störung Fahrantrieb FU 2: Überstrom / Error Drive FU 2: Überstrom'; 679 'spare / Störung Fahrantrieb FU 2: Überstrom / Error Drive FU 2: Überstrom'; 680 'spare / Störung Fahrantrieb FU 2: Überstrom / Error Drive FU 2: Überstrom'; 701 'Error hoist: FI / Störung Hubantrieb: Frequenzumrichter / Error Hoist: Frequenzumrichter'; 702 'Error hoist: spare / Störung Hubantrieb: Reserve / Error Hoist: Reserve'; 703 'Error hoist: spare / Störung Hubantrieb: Plausibilität Seilbruchschalter / Error Hoist: Plausibilität Seilbruchschalter'; 704 'Error hoist: reaches high end position / Störung Hubantrieb: Endlage oben erreicht / Error Hoist: Endlage oben erreicht'; 705 'Error hoist: reaches low end position / Störung Hubantrieb: Endlage unten erreicht / Error Hoist: Endlage unten erreicht'; 706 'Error hoist: breakage hoist rope / Störung Hubantrieb: Seilriss Hubseil / Error Hoist: Seilriss Hubseil'; 707 'Error hoist: spare / Störung Hubantrieb: Reserve / Error Hoist: Reserve'; 708 'Error hoist: spare / Störung Hubantrieb: Reserve / Error Hoist: Reserve'; 709 'Error hoist: spare / Störung Hubantrieb: Reserve / Error Hoist: Reserve'; 710 'Error hoist: spare / Störung Hubantrieb: Fangbremse und Schalter / Error Hoist: Fangbremse und Schalter'; 711 'Error hoist: spare / Störung Hubantrieb: Reserve / Error Hoist: Reserve'; 712 'Error hoist: Lowering under 500mm switch time monitoring / Störung Hubantrieb: Reserve / Error Hoist: Reserve'; 713 'Error hoist: value of encoder to high / Störung Hubantrieb: Geberwert zu hoch / Error Hoist: Geberwert zu hoch'; 714 'Error hoist: value of encoder to low / Störung Hubantrieb: Geberwert zu niedrig / Error Hoist: Geberwert zu niedrig'; 715 'Error hoist: command not plausible / Störung Hubantrieb: Hubkommando nicht plausibel / Error Hoist: Fehler Hubkommando nicht plausibel'; 716 'Error hoist: speed too high / Störung Hubantrieb: Geschwindigkeit zu hoch / Error Hoist: Geschwindigkeit zu hoch'; 717 'Error hoist: speed too low / Störung Hubantrieb: Geschwindigkeit zu niedrig / Error Hoist: Geschwindigkeit zu niedrig'; 718 'Error hoist: movement without enable / Störung Hubantrieb: Bewegung ohne Freigabe / Error Hoist: Bewegung ohne Freigabe'; 719 'Error hoist: spare / Störung Hubantrieb: Reserve / Error Hoist: Reserve'; 720 'Error hoist: jump not plausible / Störung Hubantrieb: Sprung unzulässig / Error Hoist: Sprung unzulässig'; 721 'Error hoist: movement in wrong direction / Störung Hubantrieb: Bewegung in falsche Richtung / Error Hoist: Bewegung in falsche Richtung'; 722 'Error hoist: not signal reference initiator / Störung Hubantrieb: Referenzini nicht geschaltet / Error Hoist: Referenzini nicht geschaltet'; 723 'Error hoist: signal reference initiator / Störung Hubantrieb: Referenzini nicht frei / Error Hoist: Referenzini nicht frei'; 724 'Error hoist: difference encoder to high / Störung Hubantrieb: Differenz Geberwerte zu groß / Error Hoist: Differenz Geberwerte zu groß'; 725 'Error hoist: Safety limit position reached / Störung Hubantrieb: sichere Endlage erreicht / Error Hoist: sichere Endlage erreicht'; 726 'Error hoist: no enable to lift by SDC / Störung Hubantrieb: keine Hubfreigabe vom SDC / Error Hoist: keine Hubfreigabe vom SDC'; 727 'Error hoist: spare / Störung Hubantrieb: Reserve / Error Hoist: Reserve'; 728 'Error hoist: value of rope encoder not plausible / Störung Hubantrieb: Seilgeberwert fehlerhaft / Error Hoist: Seilgeberwert fehlerhaft'; 729 'Error hoist: value of G120D not plausible / Störung Hubantrieb: G120D Positionswert fehlerhaft / Error Hoist: G120D Positionswert fehlerhaft'; 730 'Error hoist: Manipulation of encoder value, values are always the same / Störung Hubantrieb: Reserve / Error Hoist: Reserve'; 731 'Error hoist: spare / Störung Hubantrieb: Reserve / Error Hoist: Reserve'; 732 'Error hoist: spare / Störung Hubantrieb: Reserve / Error Hoist: Reserve'; 733 'Error hoist FI 1: overcurrent / Störung Hubantrieb FU 1: Überstrom / Error Hoist FU 1: Überstrom'; 734 'Error hoist FI 1: DC bus voltage overvoltage / Störung Hubantrieb FU 1: Zwischenkreisspannung Überspannung / Error Hoist FU 1: Zwischenkreisspannung Überspannung'; 735 'Error hoist FI 1: DC bus voltage undervoltage / Störung Hubantrieb FU 1: Zwischenkreisspannung Unterspannung / Error Hoist FU 1: Zwischenkreisspannung Unterspannung'; 736 'Error hoist FI 1: overtemperature / Störung Hubantrieb FU 1: Übertemperatur Kühlkörper Wechselrichter / Error Hoist FU 1: Übertemperatur Kühlkörper Wechselrichter'; 737 'Error hoist FI 1: error on driver identification / Störung Hubantrieb FU 1: Motordatenidentifikation fehlerhaft / Error Hoist FU 1: Reserve'; 738 'Error hoist FI 1: ground / Störung Hubantrieb FU 1: Erdschluss / Error Hoist FU 1: Führung durch PLC fehlt'; 739 'Error hoist FI 1: spare / Störung Hubantrieb FU 1: Reserve / Error Hoist FU 1: Reserve'; 740 'Error hoist FI 1: control requested from PLC / Störung Hubantrieb FU 1: Führung durch PLC fehlt / Error Hoist FU 1: Reserve'; 741 'Error hoist FI 1: drive overtemperature / Störung Hubantrieb FU 1: Reserve / Error Hoist FU 1: Reserve'; 742 'Error hoist FI 1: spare / Störung Hubantrieb FU 1: Reserve / Error Hoist FU 1: Reserve'; 743 'Error hoist FI 1: spare / Störung Hubantrieb FU 1: Reserve / Error Hoist FU 1: Reserve'; 744 'Error hoist FI 1: spare / Störung Hubantrieb FU 1: Reserve / Error Hoist FU 1: Reserve'; 745 'Error hoist FI 1: spare / Störung Hubantrieb FU 1: Reserve / Error Hoist FU 1: Reserve'; 746 'Error hoist FI 1: spare / Störung Hubantrieb FU 1: Reserve / Error Hoist FU 1: Reserve'; 747 'Error hoist FI 1: spare / Störung Hubantrieb FU 1: Reserve / Error Hoist FU 1: Reserve'; 748 'Error hoist FI 1: spare / Störung Hubantrieb FU 1: Reserve / Error Hoist FU 1: Führung durch PLC fehlt'; 749 'Error hoist Safety: lifting and lowering simultaneously / Störung Hubantrieb Safety: beide Drehrichtungen gleichzeitig angesteuert / Error Hoist Safety: beide Drehrichtungen gleichzeitig angesteuert'; 750 'Error hoist Safety: difference encoders to high / Störung Hubantrieb Safety: Differenz Geber 1 / 2 zu hoch / Error Hoist Safety: Differenz Geber 1 / 2 zu hoch'; 751 'Error hoist Safety: value of encoder opposite to command / Störung Hubantrieb Safety: Werte des Gebers 1 entsprechen nicht der Drehrichtung / Error Hoist Safety: Werte des Gebers 1 entsprechen nicht der Drehrichtung'; 752 'Error hoist Safety: value of G120D opposite to command / Störung Hubantrieb Safety: Werte des Gebers 2 entsprechen nicht der Drehrichtung / Error Hoist Safety: Werte des Gebers 2 entsprechen nicht der Drehrichtung'; 753 'Error hoist Safety: speed rope encoder to high / Störung Hubantrieb Safety: Geschwindigkeit Geber 1 zu hoch / Error Hoist Safety: Geschwindigkeit Geber 1 zu hoch'; 754 'Error hoist Safety: speed G120D to high / Störung Hubantrieb Safety: Geschwindigkeit Geber 2 zu hoch / Error Hoist Safety: Geschwindigkeit Geber 2 zu hoch'; 755 'Error hoist Safety: movement SLS opposite to command / Störung Hubantrieb Safety: Drehzahl des G120D entsprechen nicht der Drehrichtung / Error Hoist Safety: Drehzahl des G120D entsprechen nicht der Drehrichtung'; 756 'Error hoist Safety: speed SLS to high / Störung Hubantrieb Safety: Geschwindigkeit G120 Drehzahl zu hoch / Error Hoist Safety: Geschwindigkeit G120 Drehzahl zu hoch'; 757 'Error hoist Safety: invalid position / Störung Hubantrieb Safety: Positionswerte nicht gültig / Error Hoist Safety: Positionswerte nicht gültig'; 758 'Error hoist Safety: reference initiator not plausible / Störung Hubantrieb Safety: Referenzposition/INI nicht plausibel / Error Hoist Safety: Referenzposition/INI nicht plausibel'; 759 'Error hoist Safety: Slipping / braking distance during driver brake too high / Störung Hubantrieb Safety: Durchrutschweg/Bremsweg nach Motorhaltebremse / Error Hoist Safety: Durchrutschweg/Bremsweg nach Motorhaltebremse'; 760 'Error hoist Safety: driver holding torque not reach / Störung Hubantrieb Safety: Motorhaltemoment nicht erreicht / Error Hoist Safety: Motorhaltemoment nicht erreicht'; 761 'Error hoist Safety: feedback time catch pawl / Störung Hubantrieb Safety: Schaltzeit Hubmagnet / Error Hoist Safety: Schaltzeit Hubmagnet'; 762 'Error hoist Safety: catch pawl not plausible / Störung Hubantrieb Safety: Plausibilität von Klinkensensoren / Error Hoist Safety: Plausibilität von Klinkensensoren'; 763 'Error hoist Safety: Hoist drives in catch pawl / Störung Hubantrieb Safety: Fangklinke hat ausgelöst / Error Hoist Safety: Fangklinke hat ausgelöst'; 764 'Error hoist Safety: spare / Störung Hubantrieb Safety: Fangklinke hat ausgelöst / Error Hoist Safety: Fangklinke hat ausgelöst'; 765 'Error hoist Safety: spare / Störung Hubantrieb Safety: Fangklinke hat ausgelöst / Error Hoist Safety: Fangklinke hat ausgelöst'; 766 'Error hoist Safety: spare / Störung Hubantrieb Safety: Fangklinke hat ausgelöst / Error Hoist Safety: Fangklinke hat ausgelöst'; 767 'Error hoist Safety: spare / Störung Hubantrieb Safety: Fangklinke hat ausgelöst / Error Hoist Safety: Fangklinke hat ausgelöst'; 768 'Error hoist Safety: spare / Störung Hubantrieb Safety: Fangklinke hat ausgelöst / Error Hoist Safety: Fangklinke hat ausgelöst'; 769 'Error hoist Safety: spare / Störung Hubantrieb Safety: Fangklinke hat ausgelöst / Error Hoist Safety: Fangklinke hat ausgelöst'; 770 'Error hoist Safety: spare / Störung Hubantrieb Safety: Fangklinke hat ausgelöst / Error Hoist Safety: Fangklinke hat ausgelöst'; 771 'Error hoist Safety: spare / Störung Hubantrieb Safety: Fangklinke hat ausgelöst / Error Hoist Safety: Fangklinke hat ausgelöst'; 772 'Error hoist Safety: spare / Störung Hubantrieb Safety: Fangklinke hat ausgelöst / Error Hoist Safety: Fangklinke hat ausgelöst'; 773 'Error hoist Safety: spare / Störung Hubantrieb Safety: Fangklinke hat ausgelöst / Error Hoist Safety: Fangklinke hat ausgelöst'; 774 'Error hoist Safety: spare / Störung Hubantrieb Safety: Fangklinke hat ausgelöst / Error Hoist Safety: Fangklinke hat ausgelöst'; 775 'Error hoist Safety: spare / Störung Hubantrieb Safety: Fangklinke hat ausgelöst / Error Hoist Safety: Fangklinke hat ausgelöst'; 776 'Error hoist Safety: spare / Störung Hubantrieb Safety: Fangklinke hat ausgelöst / Error Hoist Safety: Fangklinke hat ausgelöst'; 777 'Error hoist Safety: spare / Störung Hubantrieb Safety: Fangklinke hat ausgelöst / Error Hoist Safety: Fangklinke hat ausgelöst'; 778 'Error hoist Safety: spare / Störung Hubantrieb Safety: Fangklinke hat ausgelöst / Error Hoist Safety: Fangklinke hat ausgelöst'; 779 'Error hoist Safety: spare / Störung Hubantrieb Safety: Fangklinke hat ausgelöst / Error Hoist Safety: Fangklinke hat ausgelöst'; 780 'Error hoist Safety: spare / Störung Hubantrieb Safety: Fangklinke hat ausgelöst / Error Hoist Safety: Fangklinke hat ausgelöst'; 401 'spare / Reserve'; 402 'spare / Reserve'; 403 'spare / Reserve'; 404 'spare / Reserve'; 405 'spare / Reserve'; 406 'spare / Reserve'; 407 'spare / Reserve'; 408 'spare / Reserve'; 409 'spare / Reserve'; 410 'spare / Reserve'; 411 'spare / Reserve'; 412 'spare / Reserve'; 413 'spare / Reserve'; 414 'spare / Reserve'; 415 'spare / Reserve'; 416 'spare / Reserve'; 417 'spare / Reserve'; 418 'spare / Reserve'; 419 'spare / Reserve'; 420 'spare / Reserve'; 421 'spare / Reserve'; 422 'spare / Reserve'; 423 'spare / Reserve'; 424 'spare / Reserve'; 425 'spare / Reserve'; 426 'spare / Reserve'; 427 'spare / Reserve'; 428 'spare / Reserve'; 429 'spare / Reserve'; 430 'spare / Reserve'; 431 'spare / Reserve'; 432 'spare / Reserve'; 433 'spare / Reserve'; 434 'spare / Reserve'; 435 'spare / Reserve'; 436 'spare / Reserve'; 437 'spare / Reserve'; 438 'spare / Reserve'; 439 'spare / Reserve'; 440 'spare / Reserve'; 441 'spare / Reserve'; 442 'spare / Reserve'; 443 'spare / Reserve'; 444 'spare / Reserve'; 445 'spare / Reserve'; 446 'spare / Reserve'; 447 'spare / Reserve'; 448 'spare / Reserve'; 449 'spare / Reserve'; 450 'spare / Reserve'; 451 'spare / Reserve'; 452 'spare / Reserve'; 453 'spare / Reserve'; 454 'spare / Reserve'; 455 'spare / Reserve'; 456 'spare / Reserve'; 457 'spare / Reserve'; 458 'spare / Reserve'; 459 'spare / Reserve'; 460 'spare / Reserve'; 461 'spare / Reserve'; 462 'spare / Reserve'; 463 'spare / Reserve'; 464 'spare / Reserve'; 465 'spare / Reserve'; 466 'spare / Reserve'; 467 'spare / Reserve'; 468 'spare / Reserve'; 469 'spare / Reserve'; 470 'spare / Reserve'; 471 'spare / Reserve'; 472 'spare / Reserve'; 473 'spare / Reserve'; 474 'spare / Reserve'; 475 'spare / Reserve'; 476 'spare / Reserve'; 477 'spare / Reserve'; 478 'spare / Reserve'; 479 'spare / Reserve'; 480 'spare / Reserve'; 301 'spare / Reserve'; 302 'spare / Reserve'; 303 'spare / Reserve'; 304 'spare / Reserve'; 305 'spare / Reserve'; 306 'spare / Reserve'; 307 'spare / Reserve'; 308 'spare / Reserve'; 309 'spare / Reserve'; 310 'spare / Reserve'; 311 'spare / Reserve'; 312 'spare / Reserve'; 313 'spare / Reserve'; 314 'spare / Reserve'; 315 'spare / Reserve'; 316 'spare / Reserve'; 317 'spare / Reserve'; 318 'spare / Reserve'; 319 'spare / Reserve'; 320 'spare / Reserve'; 321 'spare / Reserve'; 322 'spare / Reserve'; 323 'spare / Reserve'; 324 'spare / Reserve'; 325 'spare / Reserve'; 326 'spare / Reserve'; 327 'spare / Reserve'; 328 'spare / Reserve'; 329 'spare / Reserve'; 330 'spare / Reserve'; 331 'spare / Reserve'; 332 'spare / Reserve'; 333 'spare / Reserve / Frequency converter SPARE'; 334 'spare / Reserve / Error SPARE FC Overcurrent'; 335 'spare / Reserve / Error SPARE FC Overvoltage'; 336 'spare / Reserve / Error SPARE FC Undervoltage'; 337 'spare / Reserve / Error SPARE FC Inverter over temperature'; 338 'spare / Reserve / Error SPARE FC Motor data identification failure'; 339 'spare / Reserve / Error SPARE FC Power stack Error'; 340 'spare / Reserve / Error SPARE FC MMC contents invalid'; 341 'spare / Reserve / Error SPARE FC PLC setpoint Error'; 342 'spare / Reserve / Error SPARE FC USS setpoint Error, monitoring'; 343 'spare / Reserve / Error SPARE FC USS setpoint Error, USS master'; 344 'spare / Reserve / Error SPARE FC Errory encoder signal'; 345 'spare / Reserve / Error SPARE FC CU/PM swap'; 346 'spare / Reserve'; 347 'spare / Reserve'; 348 'spare / Reserve'; 349 'spare / Reserve'; 350 'spare / Reserve'; 351 'spare / Reserve'; 352 'spare / Reserve'; 353 'spare / Reserve'; 354 'spare / Reserve'; 355 'spare / Reserve'; 356 'spare / Reserve'; 357 'spare / Reserve'; 358 'spare / Reserve'; 359 'spare / Reserve'; 360 'spare / Reserve'; 361 'spare / Reserve'; 362 'spare / Reserve'; 363 'spare / Reserve'; 364 'spare / Reserve'; 365 'spare / Reserve / Error SPARE FC Overcurrent'; 366 'spare / Reserve / Error SPARE FC Overvoltage'; 367 'spare / Reserve / Error SPARE FC Undervoltage'; 368 'spare / Reserve / Error SPARE FC Inverter over temperature'; 369 'spare / Reserve / Error SPARE FC Motor data identification failure'; 370 'spare / Reserve / Error SPARE FC Power stack Error'; 371 'spare / Reserve / Error SPARE FC MMC contents invalid'; 372 'spare / Reserve / Error SPARE FC PLC setpoint Error'; 373 'spare / Reserve / Error SPARE FC USS setpoint Error, monitoring'; 374 'spare / Reserve / Error SPARE FC USS setpoint Error, USS master'; 375 'spare / Reserve / Error SPARE FC Errory encoder signal'; 376 'spare / Reserve / Error SPARE FC CU/PM swap'; 377 'spare / Reserve'; 378 'spare / Reserve'; 379 'spare / Reserve'; 380 'spare / Reserve'; 901 'Error SDC: spare / Reserve'; 902 'Error SDC: spare / Reserve'; 903 'Error SDC: position jump / Störung SDC Positionssprung / Error SDC Barcode Jump'; 904 'Error SDC: found no section / Störung SDC keine Sektion gefunden / Error SDC no Section found'; 905 'Error SDC: commands not plausible / Störung SDC Kommandos nicht plausibel / Error SDC wornd Commands from Main Plc'; 906 'Error SDC: position limit / Störung SDC Positionsgrenzen / Error SDC Barcode LIMIT'; 907 'Error SDC: wrong EMS no. / Störung SDC falsche EMS Nummer / Error SDC wrong EMS Number'; 908 'Error SDC: wrong section no. / Störung SDC falsche Sektion Nummer / Error SDC wrong Sektion Number'; 909 'Error SDC: spare / Reserve'; 910 'Error SDC: spare / Reserve'; 911 'Error SDC: spare / Reserve'; 912 'Error SDC: spare / Reserve'; 913 'Error SDC: spare / Reserve'; 914 'Error SDC: spare / Reserve'; 915 'Error SDC: spare / Reserve'; 916 'Error SDC: spare / Reserve'; 917 'Error SDC: communicatin with plant PLC'; 918 'Error SDC: safety communicatin with plant PLC'; 919 'Error SDC: spare'; 920 'Error SDC: spare / Reserve'; 921 'Error SDC: spare / Reserve'; 922 'Error SDC: spare / Reserve'; 923 'Error SDC: spare / Reserve'; 924 'Error SDC: spare / Reserve'

